
   // MainPos to HomePos
         AN    #IO_Button_MainPos;
         A     #Temp_IO_Status.Output.doIRBInMaintP;
         A     #Temp_IO_Status.RequestAutomatic;
         =     #Temp_IO_Status.Input.diMaintToHomeP;
   //-----
   // Cleaning MH
         A     #IO_Button_Cleaning;
         AN    #IN_FoamingCycleRunning;
         A     #Temp_IO_Status.Output.doIRBInHome;
         A     #Temp_IO_Status.RequestAutomatic;
         JCN   Cleaning;
         L     #IN_PGNO_Cleaning;
         CAW;
         T     #Temp_IO_Status.Input.GIProgNo1;
         L     0;
         T     #Temp_IO_Status.Input.GIProgNo2;
         T     #Temp_IO_Status.Input.giTeachProgNo1;
         T     #Temp_IO_Status.Input.giTeachProgNo2;
         T     #Temp_IO_Status.Input.GIMCNo;

   Cleaning:NOP   0;

         A     #IO_Button_Cleaning;
         AN    #Temp_IO_Status.Output.doIRBInHome;
         R     #IO_Button_Cleaning;

   // HomePos to CleaningPos
   // And cleaning after shot
         A     #IO_Button_Cleaning;
         A     #Temp_IO_Status.Output.doIRBInHome;
         O     #IN_CleaningRequest;
         A     #Temp_IO_Status.RequestAutomatic;
         S     #Temp_IO_Status.Input.diStartCleanMH;
   //-
         ON    #IN_MHAutomatic;
         ON    #IN_AutoStopOK;
         ON    #Temp_IO_Status.RequestAutomatic;
         O     #Temp_IO_Status.Output.doCleaningPLC;
         R     #Temp_IO_Status.Input.diStartCleanMH;
   //-----
   // Testshot MH
         A     #IO_Button_Testshot;
         AN    #IN_FoamingCycleRunning;
         A     #Temp_IO_Status.Output.doIRBInHome;
         A     #Temp_IO_Status.RequestAutomatic;
         JCN   Testshot;
         L     #IN_PGNO_Testshot;
         CAW;
         T     #Temp_IO_Status.Input.GIProgNo1;
         L     0;
         T     #Temp_IO_Status.Input.GIProgNo2;
         T     #Temp_IO_Status.Input.giTeachProgNo1;
         T     #Temp_IO_Status.Input.giTeachProgNo2;
         T     #Temp_IO_Status.Input.GIMCNo;

   Testshot:NOP   0;

         A     #IO_Button_Testshot;
         AN    #Temp_IO_Status.Output.doIRBInHome;
         R     #IO_Button_Testshot;

   // HomePos to Testshot
         A     #IO_Button_Testshot;
         AN    #Temp_IO_Status.Output.doIRBInTestP;
         A     #Temp_IO_Status.RequestAutomatic;
         =     #Temp_IO_Status.Input.diHomeToTestP;

   // Testshot to HomePos
         AN    #IO_Button_Testshot;
         A     #Temp_IO_Status.Output.doIRBInTestP;
         A     #Temp_IO_Status.RequestAutomatic;
         =     #Temp_IO_Status.Input.diTestToHomeP;

   //-----
   // Status MainPos

         L     1;
         A     #IO_Button_MainPos;
         A     #Temp_IO_Status.Output.doIRBInMaintP;
         JC    StateMainPos;

         L     3;
         A     #IO_Button_MainPos;
         AN    #Temp_IO_Status.Output.doIRBInMaintP;
         JC    StateMainPos;

         L     0;
   StateMainPos:T     #IO_State_MainPos;
   //-----
   // Status cleaning

         L     1;
   //    U     #Temp_IO_Status.Input.diStartCleanMH
         A     #Temp_IO_Status.Output.doCleaningPLC;
         JC    Statecleaning;

         L     3;
         A     #Temp_IO_Status.Input.diStartCleanMH;
         AN    #Temp_IO_Status.Output.doCleaningPLC;
         JC    Statecleaning;

         L     0;
   Statecleaning:T     #IO_State_Cleaning;
   //-----
   // Status Testshot

         L     1;
         A     #IO_Button_Testshot;
         A     #Temp_IO_Status.Output.doIRBInTestP;
         JC    Statetestshot;

         L     3;
         A     #IO_Button_Testshot;
         AN    #Temp_IO_Status.Output.doIRBInTestP;
         JC    Statetestshot;

         L     0;
   Statetestshot:T     #IO_State_Testshot;

   // for non conveyor programs the robots should not wait for the conveyor
   // Maintenance position selected robot 1
         O(;
         L     #Temp_IO_Status.Input.GIProgNo1;
         CAW;
         L     #IN_PGNO_MainPos;
         ==I;
         );
         O(;
         L     #Temp_IO_Status.Input.GIProgNo1;
         CAW;
         L     #IN_PGNO_MainPos2;
         ==I;
         );
         =     #MaintProgSel_R1;

   // MH cleaning selected robot 1
         O(;
         L     #Temp_IO_Status.Input.GIProgNo1;
         CAW;
         L     #IN_PGNO_Cleaning;
         ==I;
         );
         =     #CleanProgSel_R1;

   // MH Testshot selected robot 1
         O(;
         L     #Temp_IO_Status.Input.GIProgNo1;
         CAW;
         L     #IN_PGNO_Testshot;
         ==I;
         );
         =     #TesShotSel_R1;


   // No Program active robot 1
         O     #MaintProgSel_R1;
         O     #CleanProgSel_R1;
         O     #TesShotSel_R1;
         O(;
         L     #Temp_IO_Status.Input.GIProgNo1;
         L     #Temp_IO_Status.Input.GIProgNo2;
         OW;
         A     ==0;
         );
         A     #IN_ConfigWithTracking;
         =     #Temp_IO_Status.Input.diJumpConveyor;
END_REGION

REGION Network 8: Select automatic
         A     #Temp_IO_Status.RequestAutomatic;
   //    U     #Temp_IO_Status.Output.CMDENBL_Robot_ready
         A     #Temp_IO_Status.Output.SYSRDY_Robot_sys_ready;
         =     #Temp_IO_Status.AutomaticAccepted;
   //
         A     #Temp_IO_Status.AutomaticAccepted;
         L     S5T#2S;
         SD    #IN_TimerAutoOn;
         L     S5T#4S;
         SD    #IN_TimerAutoOnTrack;
END_REGION

REGION Network 9: Start escaping program
         A     #IN_RequestEscapeProg;
         AN    #Temp_IO_Status.Output.doCloseMouldF;
         S     #Temp_IO_Status.EscapingProgram;
         S     #Temp_IO_Status.Input.diInterrupt;
         L     S5T#3S;
         SE    #IN_TimerEscapeProg;
   //
         ON    #IN_TimerEscapeProg;
         R     #Temp_IO_Status.EscapingProgram;
         R     #Temp_IO_Status.Input.diInterrupt;
END_REGION

REGION Network 10: UOP UI 1 : IMSTP
         A     #IN_ControlVoltage;
         AN    #Temp_IO_Status.Input.diQuickStop;
         =     #Temp_IO_Status.Input.Robi_stop_extern;
END_REGION

REGION Network 11: UOP UI 3 : SFSPD
         SET;
         =     #Temp_IO_Status.Input.Robot_safety_speed;
END_REGION

REGION Network 12: UOP UI 2 : HOLD
         O(;
         O     #Temp_IO_Status.Output.Robot_Prgrun;
         O     #Temp_IO_Status.Output.Robot_Prg_paused;
         A     #Temp_IO_Status.RequestManualMode;
         A     #Temp_IO_Status.Output.SYSRDY_Robot_sys_ready;
         );
         ON    #Temp_IO_Status.Input.Robi_stop_extern;
         ON    #Temp_IO_Status.Output.SYSRDY_Robot_sys_ready;
         ON    #Temp_IO_Status.Output.CMDENBL_Robot_ready;
         A     #Temp_IO_Status.Output.do_IRB_Auto;
         NOT;
         =     #Temp_IO_Status.Input.HOLD_to_Robot;
END_REGION

REGION Network 13: UOP UI 8 : Enable robot
         SET;
         =     #Temp_IO_Status.Input.Enable_Robi_SPS_RN;
END_REGION

REGION Network 14: UOP UI 18 : Production start
   // laufendes Programm abbrechen, falls Roboter nicht im Programm ist
         A     #Temp_IO_Status.RequestAutomatic;
         AN    #Temp_IO_Status.RobotInProgram;
         A     #Temp_IO_Status.Output.Robot_Prg_paused;
         AN    #Temp_IO_Status.Output.Robot_Prgrun;
         =     #Temp_IO_Status.Input.CSTOPI_to_Robot;
   //
         A     #Temp_IO_Status.Input.PNS01;
         A     #Temp_IO_Status.RequestAutomatic;
         AN    #Temp_IO_Status.RobotInProgram;
         AN    #Temp_IO_Status.Output.Robot_Prg_paused;
         AN    #Temp_IO_Status.Output.Robot_Prgrun;
         AN    #Temp_IO_Status.Input.CSTOPI_to_Robot;
         =     #Temp_IO_Status.Input.PNS_STROBE_to_Robot;

   // Start main
         A     #IN_ControlVoltage;
         A     #Temp_IO_Status.AutomaticAccepted;
         AN    #Temp_IO_Status.RobotInProgram;
         AN    #Temp_IO_Status.Output.Robot_Prg_paused;
         =     #Temp_IO_Status.Input.PNS01;

         A     #Temp_IO_Status.Output.SNO01;  // IRB hat Nr. 1 übernommen
         AN    #Temp_IO_Status.Output.Robot_Prgrun;
         AN    #Temp_IO_Status.Input.Robot_Fault_reset;
         A     #Temp_IO_Status.RequestAutomatic;
         L     S5T#1S;  //3S
         SP    #IN_TimerStartDelay;

         A     #IN_TimerStartDelay;
         =     #Temp_IO_Status.Input.START_Robot;
   // START for CONTINUE only = FALSE, deshalb wird nur mit START_Robot gearbeitet
   //      =     #Temp_IO_Status.Input.PROD_START_to_Robot
END_REGION

REGION Network 15: Enable foamig cycle / reset / ende
         A     #IN_EnableFoamingCycle;
         AN    #IN_RequestEscapeProg;
         A     #Temp_IO_Status.AutomaticAccepted;
         =     #Temp_IO_Status.EnableFoamingCycle;
   //
         A     #Temp_IO_Status.EnableFoamingCycle;
         AN    #IN_CycleMaxWaitingTime;
         JC    spgl;
         JU    res;
END_REGION

REGION Network 16: Steps of data exchange
   spgl: L     #Temp_IO_Status.StepNumber;
   //
         JL    del;
         JU    strt;  //  0: Wait for start
         JU    wrtt;  //  1: Wait for shot times
         JU    aMld;  //  2: Number of moulds
         JU    zygo;  //  3: Start data exchange with the robot
         JU    aPr;  //  4: read program numbers
         JU    dglt;  //  5: Set data valid
         JU    dan0;  //  6: Reset data valid
         JU    Nmld;  //  7: More moulds to faom??
         JU    vpos;  //  8: wait for pre position
         JU    ssig;  //  9: foaming signals
   del:  JU    res;
   //
   res:  L     0;
         T     #Temp_IO_Status.MouldNumber;
         T     #Temp_IO_Status.OffsetForShotTime;
         T     #Temp_IO_Status.StepNumber;
         T     #Temp_IO_Status.Input.GIMCNo;
         T     #Temp_IO_Status.Input.GIProgNo1;
         T     #Temp_IO_Status.Input.GIProgNo2;
         T     #Temp_IO_Status.Input.giTeachProgNo1;
         T     #Temp_IO_Status.Input.giTeachProgNo2;
         L     1;
         T     #Temp_IO_Status.TimeNumber;
   //
         SET;
         R     #Temp_IO_Status.Input.diStartCycle;
         R     #Temp_IO_Status.Input.diReadProgNo;
         R     #Temp_IO_Status.Input.diShotDigIn;
   //
         R     #Temp_IO_Status.Input.giMouldCodeBit0;
         R     #Temp_IO_Status.Input.giMouldCodeBit1;
   //
         R     #Temp_IO_Status.StartFoamingCycle;
         R     #Temp_IO_Status.ShotTimesReceived;
         R     #Temp_IO_Status.DataTransmitted;
         R     #Temp_IO_Status.MovementProg1existing;
         R     #Temp_IO_Status.MovementProg2existing;
         R     #Temp_IO_Status.MovementProg3existing;
         R     #Temp_IO_Status.FFdoAction_01_to_Open_MH;
         R     #Temp_IO_Status.doAction_01_to_Open_MH;

         A     #Temp_IO_Status.AutomaticAccepted;
         JC    out;
         L     0;
         T     #Temp_IO_Status.RobotProgNoMould1;
         T     #Temp_IO_Status.RobotProgNoMould2;
         T     #Temp_IO_Status.RobotProgNoMould3;

         JU    out;
END_REGION

REGION Network 17: Step 0: Start foaming cycle
   strt: ON    #IN_StartPulseDataExchang;
         JC    out;

         L     #Temp_IO_Status.StepNumber;
         +     1;
         T     #Temp_IO_Status.StepNumber;
         JU    out;
END_REGION

REGION Network 18: Step 1: Wait for shot times from PUC 07
   wrtt: A(;
         O(;
         L     #Temp_IO_Status.RobotProgNoMould1;
         L     0;
         <>D;
         );
         O(;
         L     #Temp_IO_Status.RobotProgNoMould2;
         L     0;
         <>D;
         );
         O(;
         L     #Temp_IO_Status.RobotProgNoMould3;
         L     0;
         <>D;
         );
         );
         JCN   out;
   //
         L     #Temp_IO_Status.StepNumber;
         +     1;
         T     #Temp_IO_Status.StepNumber;
         JU    out;
END_REGION

REGION Network 19: Step 2: How many movement programs need to be sent
   aMld: JU    F3;
   //_________________________________________________
   // Movement for mould 3 exists
         A(;
         L     #Temp_IO_Status.RobotProgNoMould3;
         L     0;
         ==D;
         );
         JC    F2;
   //
         SET;
         S     #Temp_IO_Status.MovementProg1existing;
         S     #Temp_IO_Status.MovementProg2existing;
         S     #Temp_IO_Status.MovementProg3existing;
         S     #Temp_IO_Status.Input.giMouldCodeBit0;
         S     #Temp_IO_Status.Input.giMouldCodeBit1;
         JU    MCNr;
   //_________________________________________________
   // Movement for mould 2 exists
   F2:   O(;
         L     #Temp_IO_Status.RobotProgNoMould2;
         L     0;
         ==D;
         );
         JC    F3;
   //
         SET;
         S     #Temp_IO_Status.MovementProg1existing;
         S     #Temp_IO_Status.MovementProg2existing;
         S     #Temp_IO_Status.Input.giMouldCodeBit1;
         JU    MCNr;
   //_________________________________________________
   // Movement for mould 1 exists
   F3:   A(;
         L     #Temp_IO_Status.RobotProgNoMould1;
         L     0;
         ==I;
         );
         A(;
         L     #Temp_IO_Status.RobotProgNoMould2;
         L     0;
         ==I;
         );
         JC    MCNr;
   //
         SET;
         S     #Temp_IO_Status.MovementProg1existing;
         S     #Temp_IO_Status.Input.giMouldCodeBit0;
   //_______________________________________________
   //
   MCNr: NOP   0;
         L     #Temp_IO_Status.MCPlaceNumber;
         T     #Temp_IO_Status.Input.GIMCNo;
   //
         L     #Temp_IO_Status.StepNumber;
         +     1;
         T     #Temp_IO_Status.StepNumber;
         JU    out;
END_REGION

REGION Network 20: Step 3: Start data exchange
   zygo: NOP   0;
   //
         A     #IN_EnableDataExchange;
         S     #Temp_IO_Status.Input.diStartCycle;
         JCN   out;
   //
         L     #Temp_IO_Status.StepNumber;
         +     1;
         T     #Temp_IO_Status.StepNumber;
         JU    out;
END_REGION

REGION Network 21: Step 4: Read the actuall mould number
   aPr:  NOP   0;
   //
         A     #Temp_IO_Status.MovementProg1existing;
         JCN   a2FT;
         SET;
         R     #Temp_IO_Status.MovementProg1existing;
   //
         L     #Temp_IO_Status.RobotProgNoMould1;
         CAW;
         T     #Temp_IO_Status.Input.GIProgNo1;
         L     #Temp_IO_Status.RobotProgNoMould2;
         CAW;
         T     #Temp_IO_Status.Input.GIProgNo2;
   //
         JU    aPre;
   ///
   a2FT: A     #Temp_IO_Status.MovementProg2existing;
         JCN   a3FT;
         SET;
         R     #Temp_IO_Status.MovementProg2existing;
   //
         L     #Temp_IO_Status.RobotProgNoMould2;
         CAW;
         T     #Temp_IO_Status.Input.GIProgNo1;
   //
         JU    aPre;
   //
   a3FT: A     #Temp_IO_Status.MovementProg3existing;
         JCN   aPre;
         SET;
         R     #Temp_IO_Status.MovementProg3existing;
   //
         L     #Temp_IO_Status.RobotProgNoMould3;
         CAW;
         T     #Temp_IO_Status.Input.GIProgNo1;
   //
         JU    aPre;
   //
   aPre: L     #Temp_IO_Status.StepNumber;
         +     1;
         T     #Temp_IO_Status.StepNumber;
         JU    out;
END_REGION

REGION Network 22: Step 5: Set data valid signal
   dglt: S     #Temp_IO_Status.Input.diReadProgNo;
   //
         L     #Temp_IO_Status.StepNumber;
         +     1;
         T     #Temp_IO_Status.StepNumber;
         JU    out;
END_REGION

REGION Network 23: Step 6: reset data valid signal robot has read the information
   dan0: AN    #Temp_IO_Status.Output.doProgNoRead;
         JC    out;
         R     #Temp_IO_Status.Input.diReadProgNo;
   //
         L     #Temp_IO_Status.StepNumber;
         +     1;
         T     #Temp_IO_Status.StepNumber;
         JU    out;
END_REGION

REGION Network 24: Step 7: Wait until robot can receive new data
   Nmld: NOP   0;
   //
         A     #Temp_IO_Status.Output.doProgNoRead;
         JC    out;
   //
         AN    #Temp_IO_Status.MovementProg1existing;
         AN    #Temp_IO_Status.MovementProg2existing;
         AN    #Temp_IO_Status.MovementProg3existing;
         JC    shot;
   //
         L     4;  // 4: Next movement program
         T     #Temp_IO_Status.StepNumber;
         JU    out;
   //
   shot: L     #Temp_IO_Status.StepNumber;
         +     1;
         T     #Temp_IO_Status.StepNumber;
         JU    out;
END_REGION

REGION Network 25: Step 8: Wait until homeposition was left
   vpos: NOP   0;
         A     #Temp_IO_Status.Output.doIRBInHome;
         JC    out;
   //
         R     #Temp_IO_Status.Input.diStartCycle;

         L     0;
         T     #Temp_IO_Status.RobotProgNoMould1;
         T     #Temp_IO_Status.RobotProgNoMould2;
         T     #Temp_IO_Status.RobotProgNoMould3;

         L     #Temp_IO_Status.StepNumber;
         +     1;
         T     #Temp_IO_Status.StepNumber;
         JU    out;
END_REGION

REGION Network 26: Step 9: Wait until cycle end was sent
   ssig: NOP   0;
         A     #IN_EnableShotFromPU;
         A(;
         O     #Temp_IO_Status.Input.diShotDigIn;
         ON    #Temp_IO_Status.Output.doShotDigOut;
         );
         =     #Temp_IO_Status.Input.diShotDigIn;
   //
   // For safety reasons: open MH with ramp of the signal
   //
         A     #Temp_IO_Status.Output.doShotDigOut;
         FP    #Temp_IO_Status.FFdoAction_01_to_Open_MH;
         S     #Temp_IO_Status.doAction_01_to_Open_MH;
   //
         O     #IN_PulseShotEnd;
         ON    #IN_FoamingCycleRunning;
         ON    #Temp_IO_Status.Output.doShotDigOut;
         ON    #IN_EnableShotFromPU;
         R     #Temp_IO_Status.doAction_01_to_Open_MH;

   // End of cycle signal from robot
         AN    #Temp_IO_Status.Output.doCycleEnd;
         JC    out;
   //
         L     #Temp_IO_Status.StepNumber;
         +     1;
         T     #Temp_IO_Status.StepNumber;
         JU    out;
END_REGION

REGION Network 27: Save data
   out:  CALL  DPWR_DAT
         ( LADDR   := #IN_AdressRobIO,
           RECORD  := #Temp_IO_Status.Input,
           RET_VAL := #RetValSFC
         );

         CALL  BLKMOV
         ( SRCBLK  := #Temp_IO_Status,
           RET_VAL := #RetValSFC,
           DSTBLK  := #AnypointerStatus
         );
   //
         CALL  BLKMOV
         ( SRCBLK  := #Temp_IO_Fault,
           RET_VAL := #RetValSFC,
           DSTBLK  := #AnypointerFaults
         );
END_REGION
END_FUNCTION

FUNCTION "FC2001_KM_FRA" : Void   // FC2001, STL
TITLE = Sonderschnittstelle Faurecia Taster modifizieren
{ S7_Optimized_Access := 'TRUE' }
VERSION : 0.1
   VAR_TEMP
      Quitt : Bool;
      BildNr4 : Bool;
      Ret_Value : Int;
   END_VAR
BEGIN

REGION Network 1: Einlesen der Daten vom Koppler

         CALL  BLKMOV
         ( SRCBLK  := "FRA_KM_input",
           RET_VAL := #Ret_Value,
           DSTBLK  := "DB2000_FRA<->KM".Input
         );
END_REGION

REGION Network 2: Störungen über die Schnitsttelle quittieren

         A     "DB2000_FRA<->KM".Input.comandstatus.Reset_Fault;
         A     "S_Automatic_MH01";
         O     "T_QuitFault";
         =     "FRA_KM_Quitt";  // "T_Stoerung_quitt"
END_REGION

REGION Network 3: Watchdog Signal verarbeiten
END_REGION

REGION Network 4: Reduzierten Kreislauf einschalten üder die Schnittstelle
         A     "DB2000_FRA<->KM".Input.comandstatus.RedCirc;
         FP    "FRA_KM_HM_FP_Circulation";
         A     "S_Automatic_MH01";
         =     "FRA_KM_FP_Circulation";

         A     "FRA_KM_FP_Circulation";
         A     "DB619_State_MPart".Recirculation[1].Switch_Reduced;
         R     "DB619_State_MPart".Recirculation[1].Switch_Reduced;
         JC    g1;

         A     "FRA_KM_FP_Circulation";
         AN    "DB619_State_MPart".Recirculation[1].Switch_Reduced;
         S     "DB619_State_MPart".Recirculation[1].Switch_Reduced;

   g1:   NOP   0;
END_REGION

REGION Network 5: Service- Betrieb umschalten über die Schnittstelle
   // Service - Betrieb darf von der Schnittstelle nur geschaltet werden, wenn der 
   // Wahlschalter am MK auf Automatik steht, so dass im MK-Handbetrieb nicht von der 
   // Schnittstelle unbeabsichtigt umgeschaltet werden kann.
   // Im Bild Gruppe MK werden die [1] Variablen ständig durch [0] geschrieben
   // Und somit kommt der Befehl von FRA nicht durch
   //      L     "TP-Bereichszeiger".Picturenumber.Bildnummer
   //      L     4
   //      ==I
   //      =     #BildNr4

   //      U     "DB2000_FRA<->KM".Input.comandstatus.Service
   //      FP    "FRA_KM_HM_FP_Betrieb"
   //      U     "S_Automatic_MH01"
   //      =     "FRA_KM_FP_Betrieb"

   //      U     #BildNr4
   //      U     "DB2000_FRA<->KM".Input.comandstatus.Service
   //      U     "S_Automatic_MH01"
   //      R     "DB614_MH_State".MH_Status[0].Switch_Service_ON_OFF
   //      SPB   g2

   //      UN    #BildNr4
   //      U     "DB2000_FRA<->KM".Input.comandstatus.Service
   //      U     "S_Automatic_MH01"
   //      R     "DB614_MH_State".MH_Status[1].Switch_Service_ON_OFF
   //      SPB   g2

   //      U     #BildNr4
   //      UN    "DB2000_FRA<->KM".Input.comandstatus.Service
   //      U     "S_Automatic_MH01"
   //      S     "DB614_MH_State".MH_Status[0].Switch_Service_ON_OFF
   //      SPB   g2

   //      UN    #BildNr4
   //      UN    "DB2000_FRA<->KM".Input.comandstatus.Service
   //      U     "S_Automatic_MH01"
   //      S     "DB614_MH_State".MH_Status[1].Switch_Service_ON_OFF

   g2:   NOP   0;
END_REGION

REGION Network 6: Daten von FRA ins Prg 100 schreiben
   // Mit Strobe übernehmen
   // ACK Bit an FRA dass Strobe erkannt ist
         A     "DB009_Faults".Faults_Reset_FKT_M1;
         R     "FRA_KM_STG_Data";  // Störung Daten einlöesen
   //-----
         A     "DB2000_FRA<->KM".Output.Machinestatus.ACK;
         L     S5T#500MS;
         SD    "TM_CS_K2";

         A     "TM_CS_K2";
         R     "DB2000_FRA<->KM".Output.Machinestatus.ACK;

         A     "DB2000_FRA<->KM".Input.comandstatus.STROBE;
         FP    "FRA_KM_HM_FP_STROBE";
         A     "S_Automatic_MH01";
         S     "FRA_KM_FP_STROBE";

         A     "FRA_KM_FP_STROBE";
         AN    "DB2000_FRA<->KM".Output.Machinestatus.ACK;
         JCN   notr;

   // immer die Programmnummer 100
         L     100;
         T     "DB005_RS<->Extern".MC_Interface[1].Data_from_MC.Toolcode;
         T     "DB940_Tool_alloc_automatic".Alloc_stationTool[100];

   // Schusszeit
         L     "DB2000_FRA<->KM".Input.foaming_values.shottime;
         DTR;
         L     1000.0;
         /R;
         T     "DB925_ShotData_1".Tool[100].Shot[1].FoamingTime;

   // Durchflüsse in 0.1g/s
         L     "DB2000_FRA<->KM".Input.foaming_values.flow_C1;
         ITD;
         DTR;
         L     10.0;
         /R;
         T     "DB925_ShotData_1".Tool[100].Shot[1].Flow[1];

         L     "DB2000_FRA<->KM".Input.foaming_values.flow_C2;
         ITD;
         DTR;
         L     10.0;
         /R;
         T     "DB925_ShotData_1".Tool[100].Shot[1].Flow[2];


   // Gewicht pro Sekunde in g
         L     "DB925_ShotData_1".Tool[100].Shot[1].Flow[1];
         L     "DB925_ShotData_1".Tool[100].Shot[1].Flow[2];
         +R;
   //      T     "DB2000_FRA<->KM".AP_Weight
   //      DTR
         T     "DB925_ShotData_1".Tool[100].Shot[1].PartWeight;

   // Druck K1
         L     "DB2000_FRA<->KM".Input.foaming_values.pressure_C1;
         ITD;
         DTR;
         L     10.0;
         /R;
         T     "DB925_ShotData_1".Tool[100].Shot[1].Pressure[1];
   // Druck K2
         L     "DB2000_FRA<->KM".Input.foaming_values.pressure_C2;
         ITD;
         DTR;
         L     10.0;
         /R;
         T     "DB925_ShotData_1".Tool[100].Shot[1].Pressure[2];

   // RK
         A     "DB2000_FRA<->KM".Input.foaming_values.CP_AFTER_SHOT;
         =     "DB925_ShotData_1".Tool[100].Shot[1].CPMoveAfterShot;
   // Daten wurden gelesen
         SET;
         R     "FRA_KM_FP_STROBE";
         S     "DB930_Tools".Tool[100].EnableTool;

   // Überprüfung ob Daten Gültig
   // Wenn nicht dann Störung ausgeben!
         A(;
         L     "DB2000_FRA<->KM".Input.foaming_values.shottime;
         L     200;
         >=D;
         );
         A(;
         L     "DB2000_FRA<->KM".Input.foaming_values.flow_C1;
         L     0;
         >=I;
         );
         A(;
         L     "DB2000_FRA<->KM".Input.foaming_values.flow_C2;
         L     0;
         >=I;
         );
         NOT;
         S     "FRA_KM_STG_Data";  // Störung Daten einlöesen

         A     "FRA_KM_STG_Data";

   // ACK bit setzen, an FRA
         AN    "FRA_KM_STG_Data";  // Störung Daten einlöesen
         =     "DB2000_FRA<->KM".Output.Machinestatus.ACK;
   //-
   notr: NOP   0;
END_REGION

REGION Network 7: Signal von der Schnittstelle
   // Sie startet den Zyklus über die FT Schnittstelle 1
   // Schnittstelle stoppen
         O     "DB2000_FRA<->KM".Input.comandstatus.STOP;
         O     "S_Manuel_MH01";
         =     "DB005_RS<->Extern".MC_Interface[1].Data_from_MC.Selected;

   // Schnittstelle Starten
         A     "DB2000_FRA<->KM".Input.comandstatus.STROBE;
         A     "S_Automatic_MH01";
         S     "DB005_RS<->Extern".MC_Interface[1].Data_from_MC.Shot_preperation;

   // Mischkopf öffnen
   // Damit bei "hängendem Signal" nicht dauernd geschäumt wird vertauscht!

         O     "DB005_RS<->Extern".MC_Interface[1].Data_to_MC.Shot_end;
         ON    "DB005_RS<->Extern".MC_Interface[1].Data_from_MC.Selected;
         ON    "DB619_State_MPart".Cycle[1].Release;
         O     "DB825_Error_Interface".Interface_externalPlant[1].FLT_Watchdog;
         R     "DB005_RS<->Extern".MC_Interface[1].Data_from_MC.Shot_release;
         R     "DB005_RS<->Extern".MC_Interface[1].Data_from_MC.Shot_preperation;

         A     "DB2000_FRA<->KM".Input.comandstatus.STARTSHOT;
         A     "S_Automatic_MH01";
         S     "DB005_RS<->Extern".MC_Interface[1].Data_from_MC.Shot_release;

   // Reinigungskolben vorsteuern
         A     "DB2000_FRA<->KM".Input.comandstatus.CPFORWARD;
         A     "S_Automatic_MH01";
         =     "DB005_RS<->Extern".MC_Interface[1].Data_from_MC.CP_forward;
END_REGION

REGION Network 8: Signale an die Schnittstelle
   // Zyklus läuft
         A     "S_Automatic_MH01";
         A     "DB619_State_MPart".Cycle[1].running;
         A     "DB110_Interf_Program_M1".Status_IF[1].IF_is_on_1_Position;
         =     "DB2000_FRA<->KM".Output.Machinestatus.CYCLE_RUN;

   // Schuss läuft
         A     "S_Automatic_MH01";
         A     "DB619_State_MPart".Cycle[1].ShotRuns;
         A     "DB110_Interf_Program_M1".Status_IF[1].IF_is_on_1_Position;
         =     "DB2000_FRA<->KM".Output.Machinestatus.POURING;

   // Schussende
         A     "DB005_RS<->Extern".MC_Interface[1].Data_to_MC.Shot_end;
         =     "DB2000_FRA<->KM".Output.Machinestatus.SHOTEND;

   // Service mode
         A     "DB614_MH_State".MH_Status[1].Switch_Service_ON_OFF;
         =     "DB2000_FRA<->KM".Output.Machinestatus.SERVICE;

   // Reinigungskolben nicht hinten
         AN    "IPS_CP_MH01";
         A     "S_Automatic_MH01";
         =     "DB2000_FRA<->KM".Output.Machinestatus.CPFORWARD;

   // Ready nur nach abgelaufener Zeit ausgeben
         A     "S_Automatic_MH01";
         A     "DB110_Interf_Program_M1".Status_IF[1].IF_is_on_1_Position;
         A     "DB619_State_MPart".Cycle[1].Shotrelease;
         AN    "DB619_State_MPart".Cycle[1].ShotRuns;
         AN    "DB2000_FRA<->KM".Output.Machinestatus.ACK;
         =     "DB2000_FRA<->KM".Output.Machinestatus.READY;

   // Watchdog
         SET;
         =     "DB2000_FRA<->KM".Output.Machinestatus.Watchdog;

   // STG 1
         A     "DB009_Faults".Fault_State_Grp_1_M1;
         =     "DB2000_FRA<->KM".Output.Machinestatus.FAULTGROUP1;

   // Manual
         A     "S_Manuel_MH01";
         =     "DB2000_FRA<->KM".Output.Machinestatus.MANUAL;

   // Automatik
         A     "S_Automatic_MH01";
         A     "DB619_State_MPart".Cycle[1].Release;
         =     "DB2000_FRA<->KM".Output.Machinestatus.AUTO;

   // Startbutton an FRA
         A     "T_Start_MH01";
         =     "DB2000_FRA<->KM".Output.Machinestatus.Startbutton;

   // Kreislauf läuft
         O     "DB619_State_MPart".Recirculation[1].Reduced;
         O     "DB619_State_MPart".Recirculation[1].Lowpressure;
         O     "DB619_State_MPart".Recirculation[1].Highpressure;
         =     "DB2000_FRA<->KM".Output.Machinestatus.Kreislauf;
END_REGION

REGION Network 9: Actualwerte FRA aufbereiten
   // Menge K1
         L     "DB608_PV_Metering".Metering[1].Flow.PV_ActV.Value;
         L     10.0;
         *R;
         RND;
         T     "DB2000_FRA<->KM".Output.Act_Comp_Values.Flow_C1;
   // Menge K2
         L     "DB608_PV_Metering".Metering[2].Flow.PV_ActV.Value;
         L     10.0;
         *R;
         RND;
         T     "DB2000_FRA<->KM".Output.Act_Comp_Values.Flow_C2;

   // MVH Iso
         L     "DB2000_FRA<->KM".Output.Act_Comp_Values.Flow_C2;
         L     100;
         *D;
         L     "DB2000_FRA<->KM".Output.Act_Comp_Values.Flow_C1;
         /D;
         L     10;
         *D;
         T     "DB2000_FRA<->KM".Output.Act_Comp_Values.mixingratio;

   // Druck Pump K1
         L     "DB608_PV_Metering".Metering[1].Pressure.PV_ActV.Value;
         L     10.0;
         *R;
         RND;
         T     "DB2000_FRA<->KM".Output.Act_Comp_Values.Feedline_Pressure_C1;
   // Druck Pump K2
         L     "DB608_PV_Metering".Metering[2].Pressure.PV_ActV.Value;
         L     10.0;
         *R;
         RND;
         T     "DB2000_FRA<->KM".Output.Act_Comp_Values.Feedline_Pressure_C2;

   // Druck MH K1
         L     "DB619_State_MPart".ActMHPressureMa[1].Comp[1];
         L     10.0;
         *R;
         RND;
         T     "DB2000_FRA<->KM".Output.Act_Comp_Values.MH_Pressure_C1;
   // Druck MH K2
         L     "DB619_State_MPart".ActMHPressureMa[1].Comp[2];
         L     10.0;
         *R;
         RND;
         T     "DB2000_FRA<->KM".Output.Act_Comp_Values.MH_Pressure_C2;

   // Temp Tank K1
         L     "DB602_PV_Tank".Tank[1].Temp.PV_ActV.Value;
         L     10.0;
         *R;
         RND;
         T     "DB2000_FRA<->KM".Output.Act_Comp_Values.Tank_Temp_C1;
   // Temp Tank K2
         L     "DB602_PV_Tank".Tank[2].Temp.PV_ActV.Value;
         L     10.0;
         *R;
         RND;
         T     "DB2000_FRA<->KM".Output.Act_Comp_Values.Tank_Temp_C2;

   // Temp MH K1
         L     "DB619_State_MPart".ActMHTemperatureMa[1].Comp[1];
         L     10.0;
         *R;
         RND;
         T     "DB2000_FRA<->KM".Output.Act_Comp_Values.MH_Temp_C1;
   // Temp MH K2
         L     "DB619_State_MPart".ActMHTemperatureMa[1].Comp[2];
         L     10.0;
         *R;
         RND;
         T     "DB2000_FRA<->KM".Output.Act_Comp_Values.MH_Temp_C2;
END_REGION

REGION Network 10: letzten Schußdaten für FRA aufbereiten
   // last shot time
         L     "DB919_ShotResultMach".ShotResult_Ma[1].General.FoamingTime;
         L     1000.0;
         *R;
         RND;
         T     "DB2000_FRA<->KM".Output.Last_Shot_datas.shottime;

   // last mixingratio
         L     "DB919_ShotResultMach".ShotResult_Ma[1].Component.Comp[2].Mixingratio;
         L     10.0;
         *R;
         RND;
         T     "DB2000_FRA<->KM".Output.Last_Shot_datas.mixingratio;

   // last shot weight
         L     "DB919_ShotResultMach".ShotResult_Ma[1].General.PartWeight;
         L     10.0;
         *R;
         RND;
         T     "DB2000_FRA<->KM".Output.Last_Shot_datas.weight;

   // last flow C1
         L     "DB919_ShotResultMach".ShotResult_Ma[1].Component.Comp[1].Flow;
         L     10.0;
         *R;
         RND;
         T     "DB2000_FRA<->KM".Output.Last_Shot_datas.Flow_C1;
   // last flow C2
         L     "DB919_ShotResultMach".ShotResult_Ma[1].Component.Comp[2].Flow;
         L     10.0;
         *R;
         RND;
         T     "DB2000_FRA<->KM".Output.Last_Shot_datas.Flow_C2;

   // last pressure feedline C1
         L     "DB919_ShotResultMach".ShotResult_Ma[1].Component.Comp[1].Pressure;
         L     10.0;
         *R;
         RND;
         T     "DB2000_FRA<->KM".Output.Last_Shot_datas.Feedline_Pressure_C1;

   // last pressure MH C1
         L     "DB919_ShotResultMach".ShotResult_Ma[1].Component.Comp[1].PressureMH;
         L     10.0;
         *R;
         RND;
         T     "DB2000_FRA<->KM".Output.Last_Shot_datas.MH_Pressure_C1;


   // last pressure feedline C2
         L     "DB919_ShotResultMach".ShotResult_Ma[1].Component.Comp[2].Pressure;
         L     10.0;
         *R;
         RND;
         T     "DB2000_FRA<->KM".Output.Last_Shot_datas.Feedline_Pressure_C2;

   // last pressure MH C2
         L     "DB919_ShotResultMach".ShotResult_Ma[1].Component.Comp[2].PressureMH;
         L     10.0;
         *R;
         RND;
         T     "DB2000_FRA<->KM".Output.Last_Shot_datas.MH_Pressure_C2;


   // last temp mixhead C1
         L     "DB919_ShotResultMach".ShotResult_Ma[1].Component.Comp[1].TemperatureMH;
         L     10.0;
         *R;
         RND;
         T     "DB2000_FRA<->KM".Output.Last_Shot_datas.MH_Temp_C1;

   // last temp mixhead C2
         L     "DB919_ShotResultMach".ShotResult_Ma[1].Component.Comp[2].TemperatureMH;
         L     10.0;
         *R;
         RND;
         T     "DB2000_FRA<->KM".Output.Last_Shot_datas.MH_Temp_C2;
   //
END_REGION

REGION Network 11: Störungsbits
   // Alarme
   // n+48
         A     "DB829_Error_Machine".PouringCycle[1].FLT_OP_Mode;
         =     "DB2000_FRA<->KM".Output.Alarm_GRP1_1[8];
         A     "DB820_Error_general".Machine[1].ShotTimeTooShort;
         =     "DB2000_FRA<->KM".Output.Alarm_GRP1_1[9];
         A     "DB829_Error_Machine".SWU[1].FLT_No_SWU_selected;
         =     "DB2000_FRA<->KM".Output.Alarm_GRP1_1[10];
         A     "DB829_Error_Machine".SWU[1].FLT_Sel_SWU_not_released;
         =     "DB2000_FRA<->KM".Output.Alarm_GRP1_1[11];
         A     "DB829_Error_Machine".PouringCycle[1].FLT_Max_Shottime;
         =     "DB2000_FRA<->KM".Output.Alarm_GRP1_1[12];

         A     "DB829_Error_Machine".PouringCycle[1].FLT_WrongMixingheadNumber;
         =     "DB2000_FRA<->KM".Output.Alarm_GRP1_1[2];
         A     "DB824_Error_MH_CP".MH_Control[1].FLT_MH_dontOpen;
         =     "DB2000_FRA<->KM".Output.Alarm_GRP1_1[4];
         A     "DB824_Error_MH_CP".MH_Control[1].FLT_MH_dontClose;
         =     "DB2000_FRA<->KM".Output.Alarm_GRP1_1[5];

   // n+50
         A     "DB820_Error_general".Profibus_DP[1].Member[1];
         O     "DB820_Error_general".Profibus_DP[1].Member[2];
         O     "DB820_Error_general".Profibus_DP[1].Member[3];
         =     "DB2000_FRA<->KM".Output.Alarm_GRP1_2[15];

         A     "DB823_Error_Metering".MeteringPump[1].FLT_Max_pressure;
         =     "DB2000_FRA<->KM".Output.Alarm_GRP1_2[6];
         A     "DB823_Error_Metering".MeteringPump[2].FLT_Max_pressure;
         =     "DB2000_FRA<->KM".Output.Alarm_GRP1_2[7];

   // n+52
         A     "DB824_Error_MH_CP".Pressure[1, 1].Alarm_limit_plus;
         =     "DB2000_FRA<->KM".Output.Alarm_GRP1_3[10];
         A     "DB824_Error_MH_CP".Pressure[2, 1].Alarm_limit_plus;
         =     "DB2000_FRA<->KM".Output.Alarm_GRP1_3[11];

         A     "DB823_Error_Metering".MeteringPump[1].FLT_Min_Pressure;
         =     "DB2000_FRA<->KM".Output.Alarm_GRP1_3[0];
         A     "DB823_Error_Metering".MeteringPump[2].FLT_Min_Pressure;
         =     "DB2000_FRA<->KM".Output.Alarm_GRP1_3[1];
         A     "DB824_Error_MH_CP".Pressure[1, 1].Alarm_limit_minus;
         =     "DB2000_FRA<->KM".Output.Alarm_GRP1_3[4];
         A     "DB824_Error_MH_CP".Pressure[2, 1].Alarm_limit_minus;
         =     "DB2000_FRA<->KM".Output.Alarm_GRP1_3[5];

   // n+54
         A     "DB823_Error_Metering".MeteringPump[1].FLT_Prepressure;
         =     "DB2000_FRA<->KM".Output.Alarm_GRP1_4[10];
         A     "DB823_Error_Metering".MeteringPump[2].FLT_Prepressure;
         =     "DB2000_FRA<->KM".Output.Alarm_GRP1_4[11];

         A     "DB822_Error_Tank".Refilling_Tank[1].FLT_Min_Level;
         =     "DB2000_FRA<->KM".Output.Alarm_GRP1_4[4];
         A     "DB822_Error_Tank".Refilling_Tank[2].FLT_Min_Level;
         =     "DB2000_FRA<->KM".Output.Alarm_GRP1_4[5];

   // n+56
         A     "DB822_Error_Tank".ControllerTankTemp[1].Alarm_limit_minus;
         =     "DB2000_FRA<->KM".Output.Alarm_GRP1_5[8];
         A     "DB822_Error_Tank".ControllerTankTemp[2].Alarm_limit_minus;
         =     "DB2000_FRA<->KM".Output.Alarm_GRP1_5[9];
         A     "DB822_Error_Tank".Refilling_Tank[1].FLT_Max_Level;
         =     "DB2000_FRA<->KM".Output.Alarm_GRP1_5[14];
         A     "DB822_Error_Tank".Refilling_Tank[2].FLT_Max_Level;
         =     "DB2000_FRA<->KM".Output.Alarm_GRP1_5[15];

         A     "DB822_Error_Tank".ControllerTankTemp[1].Alarm_limit_plus;
         =     "DB2000_FRA<->KM".Output.Alarm_GRP1_5[2];
         A     "DB822_Error_Tank".ControllerTankTemp[2].Alarm_limit_plus;
         =     "DB2000_FRA<->KM".Output.Alarm_GRP1_5[3];

   // n+58
         A     "DB822_Error_Tank".Refilling_Tank[1].FLT_Max_Level_Triptray;
         =     "DB2000_FRA<->KM".Output.Alarm_GRP1_6[8];
         A     "DB822_Error_Tank".Refilling_Tank[2].FLT_Max_Level_Triptray;
         =     "DB2000_FRA<->KM".Output.Alarm_GRP1_6[9];
         A     "DB823_Error_Metering".MeteringPump[1].FLT_Tolerance_low;
         =     "DB2000_FRA<->KM".Output.Alarm_GRP1_6[12];
         A     "DB823_Error_Metering".MeteringPump[2].FLT_Tolerance_low;
         =     "DB2000_FRA<->KM".Output.Alarm_GRP1_6[13];

         A     "DB823_Error_Metering".MeteringPump[1].FLT_Tolerance_high;
         =     "DB2000_FRA<->KM".Output.Alarm_GRP1_6[0];
         A     "DB823_Error_Metering".MeteringPump[2].FLT_Tolerance_high;
         =     "DB2000_FRA<->KM".Output.Alarm_GRP1_6[1];
         A     "DB823_Error_Metering".Flow_Component[1].Alarm_limit_minus_MR;
         =     "DB2000_FRA<->KM".Output.Alarm_GRP1_6[4];
         A     "DB823_Error_Metering".Flow_Component[2].Alarm_limit_minus_MR;
         =     "DB2000_FRA<->KM".Output.Alarm_GRP1_6[5];

   // n+60
         A     "DB823_Error_Metering".Flow_Component[1].Alarm_limit_plus_MR;
         =     "DB2000_FRA<->KM".Output.Alarm_GRP1_7[8];
         A     "DB823_Error_Metering".Flow_Component[2].Alarm_limit_plus_MR;
         =     "DB2000_FRA<->KM".Output.Alarm_GRP1_7[9];
         A     "DB821_Error_Hydraulic".MH_Hydraulic[1].FLT_Motorprotection;
         =     "DB2000_FRA<->KM".Output.Alarm_GRP1_7[12];
         A     "DB821_Error_Hydraulic".MH_Hydraulic[1].FLT_C_Max;
         =     "DB2000_FRA<->KM".Output.Alarm_GRP1_7[13];
         A     "DB821_Error_Hydraulic".MH_Hydraulic[1].FLT_Min_Level;
         =     "DB2000_FRA<->KM".Output.Alarm_GRP1_7[14];
         A     "DB821_Error_Hydraulic".MH_Hydraulic[1].FLT_P_Max;
         =     "DB2000_FRA<->KM".Output.Alarm_GRP1_7[15];

         A     "DB823_Error_Metering".MeteringPump[1].FLT_Motorprotection;
         =     "DB2000_FRA<->KM".Output.Alarm_GRP1_7[6];
         A     "DB823_Error_Metering".MeteringPump[2].FLT_Motorprotection;
         =     "DB2000_FRA<->KM".Output.Alarm_GRP1_7[7];

   // n+62
         A     "DB824_Error_MH_CP".Temperature[1, 1].Alarm_limit_minus;
         =     "DB2000_FRA<->KM".Output.Alarm_GRP1_8[10];
         A     "DB824_Error_MH_CP".Temperature[2, 1].Alarm_limit_minus;
         =     "DB2000_FRA<->KM".Output.Alarm_GRP1_8[11];

         A     "DB823_Error_Metering".MeteringPump[1].FLT_F_converter;
         =     "DB2000_FRA<->KM".Output.Alarm_GRP1_8[0];
         A     "DB823_Error_Metering".MeteringPump[2].FLT_F_converter;
         =     "DB2000_FRA<->KM".Output.Alarm_GRP1_8[1];
         A     "DB824_Error_MH_CP".Temperature[1, 1].Alarm_limit_plus;
         =     "DB2000_FRA<->KM".Output.Alarm_GRP1_8[4];
         A     "DB824_Error_MH_CP".Temperature[2, 1].Alarm_limit_plus;
         =     "DB2000_FRA<->KM".Output.Alarm_GRP1_8[5];

   // n+66
         A     "DB823_Error_Metering".FeedPump[1].FLT_Motorprotection;
         =     "DB2000_FRA<->KM".Output.Alarm_GRP1_10[14];
         A     "DB823_Error_Metering".FeedPump[2].FLT_Motorprotection;
         =     "DB2000_FRA<->KM".Output.Alarm_GRP1_10[15];

   // n+68
         A     "DB823_Error_Metering".MeteringPump[1].FLT_Prepressure;
         =     "DB2000_FRA<->KM".Output.Alarm_GRP1_11[2];
         A     "DB823_Error_Metering".MeteringPump[2].FLT_Prepressure;
         =     "DB2000_FRA<->KM".Output.Alarm_GRP1_11[3];

   // Warnungen
   // n+80
         A     "DB822_Error_Tank".Refilling_Tank[1].FLT_Min_Level_Cycle;
         =     "DB2000_FRA<->KM".Output.Alarm_GRP2_1[12];
         A     "DB822_Error_Tank".Refilling_Tank[2].FLT_Min_Level_Cycle;
         =     "DB2000_FRA<->KM".Output.Alarm_GRP2_1[13];

   // n+84
         A     "DB821_Error_Hydraulic".MH_Hydraulic[1].FLT_WRN_C_Max;
         =     "DB2000_FRA<->KM".Output.Alarm_GRP2_3[10];

   // Meldungen
   // n+88
         A     "DB822_Error_Tank".Agitator[1].FLT_Motorprotection;
         =     "DB2000_FRA<->KM".Output.Alarm_GRP3_1[8];
         A     "DB822_Error_Tank".Agitator[2].FLT_Motorprotection;
         =     "DB2000_FRA<->KM".Output.Alarm_GRP3_1[9];

         A     "DB822_Error_Tank".Agitator[1].FLT_FrequencyConverter;
         =     "DB2000_FRA<->KM".Output.Alarm_GRP3_1[2];
         A     "DB822_Error_Tank".Agitator[2].FLT_FrequencyConverter;
         =     "DB2000_FRA<->KM".Output.Alarm_GRP3_1[3];

   // n+90
         A     "DB822_Error_Tank".Refilling_Tank[1].FLT_Fillingtime_to_long;
         =     "DB2000_FRA<->KM".Output.Alarm_GRP3_2[12];
         A     "DB822_Error_Tank".Refilling_Tank[2].FLT_Fillingtime_to_long;
         =     "DB2000_FRA<->KM".Output.Alarm_GRP3_2[13];

         A     "DB822_Error_Tank".Refilling_Tank[1].FLT_LevelSensor_broken_wire;
         =     "DB2000_FRA<->KM".Output.Alarm_GRP3_2[0];
         A     "DB822_Error_Tank".Refilling_Tank[2].FLT_LevelSensor_broken_wire;
         =     "DB2000_FRA<->KM".Output.Alarm_GRP3_2[1];

   // n+92
         A     "DB823_Error_Metering".EdgeFilter[1].FLT_Motorprotection;
         =     "DB2000_FRA<->KM".Output.Alarm_GRP3_3[0];
         A     "DB823_Error_Metering".EdgeFilter[2].FLT_Motorprotection;
         =     "DB2000_FRA<->KM".Output.Alarm_GRP3_3[1];

   // n+94
         A     "DB821_Error_Hydraulic".MH_Hydraulic[1].FLT_Filter_backflow;
         =     "DB2000_FRA<->KM".Output.Alarm_GRP3_4[10];
         A     "DB821_Error_Hydraulic".MH_Hydraulic[1].FLT_Filter_HP;
         =     "DB2000_FRA<->KM".Output.Alarm_GRP3_4[11];

   // n+96
         A     "DB829_Error_Machine".PouringCycle[1].FLT_KLZ_0;
         =     "DB2000_FRA<->KM".Output.Alarm_GRP3_5[14];
         A     "DB829_Error_Machine".PouringCycle[1].FLT_Max_Waittime;
         =     "DB2000_FRA<->KM".Output.Alarm_GRP3_5[15];

         A     "DB820_Error_general".Machine[1].Fuse_broken;
         =     "DB2000_FRA<->KM".Output.Alarm_GRP3_5[2];
         A     "DB820_Error_general".Machine[1].Air_dryer;
         =     "DB2000_FRA<->KM".Output.Alarm_GRP3_5[3];

   // n+120
         A     "DB823_Error_Metering".MeteringPump[1].FLT_FlowSDATimeOut;
         O     "DB823_Error_Metering".MeteringPump[2].FLT_FlowSDATimeOut;
         =     "DB2000_FRA<->KM".Output.Alarm_GRP3_17[10];

         A     "DB824_Error_MH_CP".Pressure[1, 1].Warning_limit_minus;
         =     "DB2000_FRA<->KM".Output.Alarm_GRP3_17[5];
         A     "DB824_Error_MH_CP".Pressure[2, 1].Warning_limit_minus;
         =     "DB2000_FRA<->KM".Output.Alarm_GRP3_17[6];

   // n+122
         A     "DB824_Error_MH_CP".Pressure[1, 1].Warning_limit_plus;
         =     "DB2000_FRA<->KM".Output.Alarm_GRP3_18[9];
         A     "DB824_Error_MH_CP".Pressure[2, 1].Warning_limit_plus;
         =     "DB2000_FRA<->KM".Output.Alarm_GRP3_18[10];
         A     "DB824_Error_MH_CP".Temperature[1, 1].Warning_limit_minus;
         =     "DB2000_FRA<->KM".Output.Alarm_GRP3_18[13];
         A     "DB824_Error_MH_CP".Temperature[2, 1].Warning_limit_minus;
         =     "DB2000_FRA<->KM".Output.Alarm_GRP3_18[14];

         A     "DB824_Error_MH_CP".Temperature[1, 1].Warning_limit_plus;
         =     "DB2000_FRA<->KM".Output.Alarm_GRP3_18[1];
         A     "DB824_Error_MH_CP".Temperature[2, 1].Warning_limit_plus;
         =     "DB2000_FRA<->KM".Output.Alarm_GRP3_18[2];
         A     "DB823_Error_Metering".Flow_Component[1].Warning_limit_minus;
         =     "DB2000_FRA<->KM".Output.Alarm_GRP3_18[5];
         A     "DB823_Error_Metering".Flow_Component[2].Warning_limit_minus;
         =     "DB2000_FRA<->KM".Output.Alarm_GRP3_18[6];

   // n+124
         A     "DB823_Error_Metering".Flow_Component[1].Warning_limit_plus;
         =     "DB2000_FRA<->KM".Output.Alarm_GRP3_19[9];
         A     "DB823_Error_Metering".Flow_Component[2].Warning_limit_plus;
         =     "DB2000_FRA<->KM".Output.Alarm_GRP3_19[10];
         A     "DB823_Error_Metering".Flow_Component[1].Warning_limit_minus_MR;
         =     "DB2000_FRA<->KM".Output.Alarm_GRP3_19[13];
         A     "DB823_Error_Metering".Flow_Component[2].Warning_limit_minus_MR;
         =     "DB2000_FRA<->KM".Output.Alarm_GRP3_19[14];

         A     "DB823_Error_Metering".Flow_Component[1].Warning_limit_plus_MR;
         =     "DB2000_FRA<->KM".Output.Alarm_GRP3_19[1];
         A     "DB823_Error_Metering".Flow_Component[2].Warning_limit_plus_MR;
         =     "DB2000_FRA<->KM".Output.Alarm_GRP3_19[2];
         A     "DB824_Error_MH_CP".MH_Control[1].WRN_ShotTimeShort;
         =     "DB2000_FRA<->KM".Output.Alarm_GRP3_19[5];
         A     "DB824_Error_MH_CP".MH_Control[1].WRN_ShotTimeLong;
         =     "DB2000_FRA<->KM".Output.Alarm_GRP3_19[6];

   // n+126
         A     "DB822_Error_Tank".ControllerTankTemp[1].Warning_limit_minus;
         =     "DB2000_FRA<->KM".Output.Alarm_GRP3_20[9];
         A     "DB822_Error_Tank".ControllerTankTemp[2].Warning_limit_minus;
         =     "DB2000_FRA<->KM".Output.Alarm_GRP3_20[10];
         A     "DB822_Error_Tank".ControllerTankTemp[1].Warning_limit_plus;
         =     "DB2000_FRA<->KM".Output.Alarm_GRP3_20[13];
         A     "DB822_Error_Tank".ControllerTankTemp[2].Warning_limit_plus;
         =     "DB2000_FRA<->KM".Output.Alarm_GRP3_20[14];

   // Not-Aus
   // n+144
         A     "DB820_Error_general".Machine[1].Controlvoltage;
         =     "DB2000_FRA<->KM".Output.Message_1[8];
         A     "DB822_Error_Tank".InterfaceContainer.FLT_containerstation;
         =     "DB2000_FRA<->KM".Output.Message_1[9];
         A     "DB820_Error_general".Machine[1].EmergencyStop.Machine;
         =     "DB2000_FRA<->KM".Output.Message_1[10];
         A     "DB820_Error_general".Machine[1].EmergencyStop.MH_Cleaner_2;
         =     "DB2000_FRA<->KM".Output.Message_1[13];

         A     "DB820_Error_general".Machine[1].EmergencyStop.External_Plant_1;
         =     "DB2000_FRA<->KM".Output.Alarm_GRP1_2[13];
   // n+146
         A     "DB822_Error_Tank".InterfaceContainer.MSG_EScontainerstation;
         =     "DB2000_FRA<->KM".Output.Message_2[6];

   // n+148
         A     "DB123_MH_IO_Signals".MH[1].IN.MH_EmergencyStop;
         =     "DB2000_FRA<->KM".Output.Message_3[8];

   // n+154
         A     "DB820_Error_general".Machine[1].Weekend_Mode;
         =     "DB2000_FRA<->KM".Output.Message_6[15];

   // n+160
         A     "DB823_Error_Metering".MeteringPump[1].Mes_StartUpDelayFU;
         =     "DB2000_FRA<->KM".Output.Message_9[11];
END_REGION

REGION Network 12: Daten auf BUS (an FRA)
   // Bits, Istwerte, Schussdaten, Reserve

         CALL  BLKMOV
         ( SRCBLK  := "DB2000_FRA<->KM".Output,
           RET_VAL := #Ret_Value,
           DSTBLK  := "FRA_KM_output"
         );
END_REGION
END_FUNCTION

FUNCTION "FC2170_TimeHandle" : Void   // FC2170, STL
{ S7_Optimized_Access := 'FALSE' }
AUTHOR : KT242
VERSION : 0.1
// Uhrzeit des AG stellen, dann an TP transferiern
   VAR_TEMP
      date_time_new : Date_And_Time;
      sfc0_ret : Int;
      sfc1_ret : Int;
      Date_new : Date;
      Time_new : Time_Of_Day;
      RetValSFC : Int;
   END_VAR
BEGIN

REGION Network 1: CPU Zeit ständig lesen
   // MP holt sich diese selbsständig alle 3600 Sekunden.
   // Datum und Uhrzeit holen
         CALL  RD_SYS_T
         ( RET_VAL := #RetValSFC,
           OUT     := "TP-Bereichszeiger".Date_Time.ActTime
         );
END_REGION

REGION Network 2: Uhrzeit stellen am TP und Übertrag an CPU
         AN    "TP-Bereichszeiger".Date_Time.Start_AG_Transfer;  // Startbit, beim Drücken von Speichern im OP
         BEC;
END_REGION

REGION Network 3: Uhr am AG stellen
         CALL  WR_SYS_T
         ( IN      := "TP-Bereichszeiger".Date_Time.SetTime,
           RET_VAL := #sfc0_ret
         );

         SET;
         R     "TP-Bereichszeiger".Date_Time.Start_AG_Transfer;  // Startbit reseten

         BEU;
END_REGION
END_FUNCTION

FUNCTION "PartCounter" : Void   // FC5001, SCL
{ S7_Optimized_Access := 'FALSE' }
VERSION : 0.1
   VAR_TEMP
      i : Int;
   END_VAR
BEGIN

